screen "Dev_DO_2" 800x480, template "Settings"
   TextField "Text field_4" at 134,11 size 130x26; Text 'выход 1'
   TextField "Text field_5" at 286,11 size 130x26; Text 'выход 2'
   TextField "Text field_29" at 438,11 size 130x26; Text 'выход 3'
   TextField "Text field_33" at 590,11 size 130x26; Text 'выход 4'
   TextField "Text field_17" at 134,283 size 130x26; Text 'выход 9'
   TextField "Text field_25" at 286,283 size 130x26; Text 'выход 10'
   TextField "Text field_9" at 134,147 size 130x26; Text 'выход 5'
   TextField "Text field_13" at 286,147 size 130x26; Text 'выход 6'
   TextField "Text field_21" at 438,147 size 130x26; Text 'выход 7'
   TextField "Text field_41" at 590,147 size 130x26; Text 'выход 8'
   TextField "Text field_37" at 590,283 size 130x26; Text 'выход 12'
   Button "Button_2" at 134,40 size 130x22; TextOff 'Авто'; Authorization "Operate"; TextList "Hand"
      on Click: InvertBit("DOx_Hand_x_1")
      Appearance <- "DOx_Hand_x_1"
      ProcessValue <- "DOx_Hand_x_1"
   Button "Button_13" at 134,65 size 60x20; TextOff 'Вкл'; Authorization "Operate"
      on Click: SetBit("DOx_Start_M_x_1")
      Appearance <- "DOx_Start_M_x_1"
   Button "Button_26" at 244,89 size 20x20; TextOff 'Text'; Authorization "User administration"; PictureList "ok_green"
      on Click: InvertBit("DOx_Inverse_x_1")
      ProcessValue <- "DOx_Inverse_x_1"
   TextField "Text field_1" at 133,85 size 91x23; Text 'Инверсия:'
   IOField "I/O field_1" at 176,109 size 30x24; Authorization "Developer"; FormatPattern 99
      ProcessValue <- "DOx_ADDR_Byte_x_1"
   IOField "I/O field_2" at 216,109 size 20x24; Authorization "Developer"; FormatPattern 9
      ProcessValue <- "DOx_ADDR_Bit_x_1"
   TextField "Text field_2" at 158,109 size 20x23; Text 'Q'
   TextField "Text field_3" at 205,109 size 13x23; Text '.'
   Button "Button_1" at 286,40 size 130x22; TextOff 'Авто'; Authorization "Operate"; TextList "Hand"
      on Click: InvertBit("DOx_Hand_x_2")
      Appearance <- "DOx_Hand_x_2"
      ProcessValue <- "DOx_Hand_x_2"
   Button "Button_5" at 286,65 size 60x20; TextOff 'Вкл'; Authorization "Operate"
      on Click: SetBit("DOx_Start_M_x_2")
      Appearance <- "DOx_Start_M_x_2"
   Button "Button_6" at 396,89 size 20x20; TextOff 'Text'; PictureList "ok_green"; Authorization "User administration"
      on Click: InvertBit("DOx_Inverse_x_2")
      ProcessValue <- "DOx_Inverse_x_2"
   TextField "Text field_6" at 285,85 size 91x23; Text 'Инверсия:'
   IOField "I/O field_3" at 328,109 size 30x24; Authorization "Developer"; FormatPattern 99
      ProcessValue <- "DOx_ADDR_Byte_x_2"
   IOField "I/O field_4" at 368,109 size 20x24; Authorization "Developer"; FormatPattern 9
      ProcessValue <- "DOx_ADDR_Bit_x_2"
   TextField "Text field_7" at 310,109 size 20x23; Text 'Q'
   TextField "Text field_8" at 357,109 size 13x23; Text '.'
   Button "Button_29" at 438,40 size 130x22; TextOff 'Авто'; Authorization "Operate"; TextList "Hand"
      on Click: InvertBit("DOx_Hand_x_3")
      Appearance <- "DOx_Hand_x_3"
      ProcessValue <- "DOx_Hand_x_3"
   Button "Button_31" at 438,65 size 60x20; TextOff 'Вкл'; Authorization "Operate"
      on Click: SetBit("DOx_Start_M_x_3")
      Appearance <- "DOx_Start_M_x_3"
   Button "Button_32" at 548,89 size 20x20; TextOff 'Text'; PictureList "ok_green"; Authorization "User administration"
      on Click: InvertBit("DOx_Inverse_x_3")
      ProcessValue <- "DOx_Inverse_x_3"
   TextField "Text field_30" at 437,85 size 91x23; Text 'Инверсия:'
   IOField "I/O field_15" at 480,109 size 30x24; Authorization "Developer"; FormatPattern 99
      ProcessValue <- "DOx_ADDR_Byte_x_3"
   IOField "I/O field_16" at 520,109 size 20x24; Authorization "Developer"; FormatPattern 9
      ProcessValue <- "DOx_ADDR_Bit_x_3"
   TextField "Text field_31" at 462,109 size 20x23; Text 'Q'
   TextField "Text field_32" at 509,109 size 13x23; Text '.'
   Button "Button_33" at 590,40 size 130x22; TextOff 'Авто'; Authorization "Operate"; TextList "Hand"
      on Click: InvertBit("DOx_Hand_x_4")
      Appearance <- "DOx_Hand_x_4"
      ProcessValue <- "DOx_Hand_x_4"
   Button "Button_35" at 590,65 size 60x20; TextOff 'Вкл'; Authorization "Operate"
      on Click: SetBit("DOx_Start_M_x_4")
      Appearance <- "DOx_Start_M_x_4"
   Button "Button_36" at 700,89 size 20x20; TextOff 'Text'; PictureList "ok_green"; Authorization "User administration"
      on Click: InvertBit("DOx_Inverse_x_4")
      ProcessValue <- "DOx_Inverse_x_4"
   TextField "Text field_34" at 589,85 size 91x23; Text 'Инверсия:'
   IOField "I/O field_17" at 632,109 size 30x24; Authorization "Developer"; FormatPattern 99
      ProcessValue <- "DOx_ADDR_Byte_x_4"
   IOField "I/O field_18" at 672,109 size 20x24; Authorization "Developer"; FormatPattern 9
      ProcessValue <- "DOx_ADDR_Bit_x_4"
   TextField "Text field_35" at 614,109 size 20x23; Text 'Q'
   TextField "Text field_36" at 661,109 size 13x23; Text '.'
   Button "Button_7" at 134,176 size 130x22; TextOff 'Авто'; Authorization "Operate"; TextList "Hand"
      on Click: InvertBit("DOx_Hand_x_5")
      Appearance <- "DOx_Hand_x_5"
      ProcessValue <- "DOx_Hand_x_5"
   Button "Button_9" at 134,201 size 60x20; TextOff 'Вкл'; Authorization "Operate"
      on Click: SetBit("DOx_Start_M_x_5")
      Appearance <- "DOx_Start_M_x_5"
   Button "Button_10" at 244,225 size 20x20; TextOff 'Text'; PictureList "ok_green"; Authorization "User administration"
      on Click: InvertBit("DOx_Inverse_x_5")
      ProcessValue <- "DOx_Inverse_x_5"
   TextField "Text field_10" at 133,221 size 91x23; Text 'Инверсия:'
   IOField "I/O field_5" at 176,245 size 30x24; Authorization "Developer"; FormatPattern 99
      ProcessValue <- "DOx_ADDR_Byte_x_5"
   IOField "I/O field_6" at 216,245 size 20x24; Authorization "Developer"; FormatPattern 9
      ProcessValue <- "DOx_ADDR_Bit_x_5"
   TextField "Text field_11" at 158,245 size 20x23; Text 'Q'
   TextField "Text field_12" at 205,245 size 13x23; Text '.'
   Button "Button_11" at 286,176 size 130x22; TextOff 'Авто'; Authorization "Operate"; TextList "Hand"
      on Click: InvertBit("DOx_Hand_x_6")
      Appearance <- "DOx_Hand_x_6"
      ProcessValue <- "DOx_Hand_x_6"
   Button "Button_14" at 286,201 size 60x20; TextOff 'Вкл'; Authorization "Operate"
      on Click: SetBit("DOx_Start_M_x_6")
      Appearance <- "DOx_Start_M_x_6"
   Button "Button_15" at 396,225 size 20x20; TextOff 'Text'; Authorization "User administration"; PictureList "ok_green"
      on Click: InvertBit("DOx_Inverse_x_6")
      ProcessValue <- "DOx_Inverse_x_6"
   TextField "Text field_14" at 285,221 size 91x23; Text 'Инверсия:'
   IOField "I/O field_7" at 328,245 size 30x24; Authorization "Developer"; FormatPattern 99
      ProcessValue <- "DOx_ADDR_Byte_x_6"
   IOField "I/O field_8" at 368,245 size 20x24; Authorization "Developer"; FormatPattern 9
      ProcessValue <- "DOx_ADDR_Bit_x_6"
   TextField "Text field_15" at 310,245 size 20x23; Text 'Q'
   TextField "Text field_16" at 357,245 size 13x23; Text '.'
   Button "Button_20" at 438,176 size 130x22; TextOff 'Авто'; Authorization "Operate"; TextList "Hand"
      on Click: InvertBit("DOx_Hand_x_7")
      Appearance <- "DOx_Hand_x_7"
      ProcessValue <- "DOx_Hand_x_7"
   Button "Button_22" at 438,201 size 60x20; TextOff 'Вкл'; Authorization "Operate"
      on Click: SetBit("DOx_Start_M_x_7")
      Appearance <- "DOx_Start_M_x_7"
   Button "Button_23" at 548,225 size 20x20; TextOff 'Text'; Authorization "User administration"; PictureList "ok_green"
      on Click: InvertBit("DOx_Inverse_x_7")
      ProcessValue <- "DOx_Inverse_x_7"
   TextField "Text field_22" at 437,221 size 91x23; Text 'Инверсия:'
   IOField "I/O field_11" at 480,245 size 30x24; Authorization "Developer"; FormatPattern 99
      ProcessValue <- "DOx_ADDR_Byte_x_7"
   IOField "I/O field_12" at 520,245 size 20x24; Authorization "Developer"; FormatPattern 9
      ProcessValue <- "DOx_ADDR_Bit_x_7"
   TextField "Text field_23" at 462,245 size 20x23; Text 'Q'
   TextField "Text field_24" at 509,245 size 13x23; Text '.'
   Button "Button_41" at 590,176 size 130x22; TextOff 'Авто'; Authorization "Operate"; TextList "Hand"
      on Click: InvertBit("DOx_Hand_x_8")
      Appearance <- "DOx_Hand_x_8"
      ProcessValue <- "DOx_Hand_x_8"
   Button "Button_43" at 590,201 size 60x20; TextOff 'Вкл'; Authorization "Operate"
      on Click: SetBit("DOx_Start_M_x_8")
      Appearance <- "DOx_Start_M_x_8"
   Button "Button_44" at 700,225 size 20x20; TextOff 'Text'; Authorization "User administration"; PictureList "ok_green"
      on Click: InvertBit("DOx_Inverse_x_8")
      ProcessValue <- "DOx_Inverse_x_8"
   TextField "Text field_42" at 589,221 size 91x23; Text 'Инверсия:'
   IOField "I/O field_21" at 632,245 size 30x24; Authorization "Developer"; FormatPattern 99
      ProcessValue <- "DOx_ADDR_Byte_x_8"
   IOField "I/O field_22" at 672,245 size 20x24; Authorization "Developer"; FormatPattern 9
      ProcessValue <- "DOx_ADDR_Bit_x_8"
   TextField "Text field_43" at 614,245 size 20x23; Text 'Q'
   TextField "Text field_44" at 661,245 size 13x23; Text '.'
   Button "Button_24" at 134,312 size 130x22; TextOff 'Авто'; Authorization "Operate"; TextList "Hand"
      on Click: InvertBit("DOx_Hand_x_9")
      Appearance <- "DOx_Hand_x_9"
      ProcessValue <- "DOx_Hand_x_9"
   Button "Button_27" at 134,337 size 60x20; TextOff 'Вкл'; Authorization "Operate"
      on Click: SetBit("DOx_Start_M_x_9")
      Appearance <- "DOx_Start_M_x_9"
   Button "Button_28" at 244,361 size 20x20; TextOff 'Text'; PictureList "ok_green"; Authorization "User administration"
      on Click: InvertBit("DOx_Inverse_x_9")
      ProcessValue <- "DOx_Inverse_x_9"
   TextField "Text field_18" at 133,357 size 91x23; Text 'Инверсия:'
   IOField "I/O field_9" at 176,381 size 30x24; Authorization "Developer"; FormatPattern 99
      ProcessValue <- "DOx_ADDR_Byte_x_9"
   IOField "I/O field_10" at 216,381 size 20x24; Authorization "Developer"; FormatPattern 9
      ProcessValue <- "DOx_ADDR_Bit_x_9"
   TextField "Text field_19" at 158,381 size 20x23; Text 'Q'
   TextField "Text field_20" at 205,381 size 13x23; Text '.'
   Button "Button_37" at 286,312 size 130x22; TextOff 'Авто'; Authorization "Operate"; TextList "Hand"
      on Click: InvertBit("DOx_Hand_x_10")
      Appearance <- "DOx_Hand_x_10"
      ProcessValue <- "DOx_Hand_x_10"
   Button "Button_39" at 286,337 size 60x20; TextOff 'Вкл'; Authorization "Operate"
      on Click: SetBit("DOx_Start_M_x_10")
      Appearance <- "DOx_Start_M_x_10"
   Button "Button_40" at 396,361 size 20x20; TextOff 'Text'; Authorization "User administration"; PictureList "ok_green"
      on Click: InvertBit("DOx_Inverse_x_10")
      ProcessValue <- "DOx_Inverse_x_10"
   TextField "Text field_26" at 285,357 size 91x23; Text 'Инверсия:'
   IOField "I/O field_13" at 328,381 size 30x24; Authorization "Developer"; FormatPattern 99
      ProcessValue <- "DOx_ADDR_Byte_x_10"
   IOField "I/O field_14" at 368,381 size 20x24; Authorization "Developer"; FormatPattern 9
      ProcessValue <- "DOx_ADDR_Bit_x_10"
   TextField "Text field_27" at 310,381 size 20x23; Text 'Q'
   TextField "Text field_28" at 357,381 size 13x23; Text '.'
   Button "Button_48" at 590,312 size 130x22; TextOff 'Авто'; Authorization "Operate"; TextList "Hand"
      on Click: InvertBit("DOx_Hand_x_12")
      Appearance <- "DOx_Hand_x_12"
      ProcessValue <- "DOx_Hand_x_12"
   Button "Button_50" at 590,337 size 60x20; TextOff 'Вкл'; Authorization "Operate"
      on Click: SetBit("DOx_Start_M_x_12")
      Appearance <- "DOx_Start_M_x_12"
   Button "Button_51" at 700,361 size 20x20; TextOff 'Text'; Authorization "User administration"; PictureList "ok_green"
      on Click: InvertBit("DOx_Inverse_x_12")
      ProcessValue <- "DOx_Inverse_x_12"
   TextField "Text field_45" at 589,357 size 91x23; Text 'Инверсия:'
   IOField "I/O field_23" at 632,381 size 30x24; Authorization "Developer"; FormatPattern 99
      ProcessValue <- "DOx_ADDR_Byte_x_12"
   IOField "I/O field_24" at 672,381 size 20x24; Authorization "Developer"; FormatPattern 9
      ProcessValue <- "DOx_ADDR_Bit_x_12"
   TextField "Text field_46" at 614,381 size 20x23; Text 'Q'
   TextField "Text field_47" at 661,381 size 13x23; Text '.'
   TextField "Text field_38" at 438,283 size 130x26; Text 'выход 11'
   Button "Button_45" at 438,312 size 130x22; TextOff 'Авто'; Authorization "Operate"; TextList "Hand"
      on Click: InvertBit("DOx_Hand_x_11")
      Appearance <- "DOx_Hand_x_11"
      ProcessValue <- "DOx_Hand_x_11"
   Button "Button_47" at 438,337 size 60x20; TextOff 'Вкл'; Authorization "Operate"
      on Click: SetBit("DOx_Start_M_x_11")
      Appearance <- "DOx_Start_M_x_11"
   Button "Button_52" at 548,361 size 20x20; TextOff 'Text'; PictureList "ok_green"; Authorization "User administration"
      on Click: InvertBit("DOx_Inverse_x_11")
      ProcessValue <- "DOx_Inverse_x_11"
   TextField "Text field_39" at 437,357 size 91x23; Text 'Инверсия:'
   IOField "I/O field_19" at 480,381 size 30x24; Authorization "Developer"; FormatPattern 99
      ProcessValue <- "DOx_ADDR_Byte_x_11"
   IOField "I/O field_20" at 520,381 size 20x24; Authorization "Developer"; FormatPattern 9
      ProcessValue <- "DOx_ADDR_Bit_x_11"
   TextField "Text field_40" at 462,381 size 20x23; Text 'Q'
   TextField "Text field_48" at 509,381 size 13x23; Text '.'
   Button "Button_16" at 128,440 size 75x30; TextOff 'Стр.1'; Authorization "Operate"
      on Click: SetTag("DOx", 210); ActivateScreen("Dev_DI_1", 0)
      Visibility <- "Support_DB_All_DOs"
      Appearance <- "DOx"
   Button "Button_17" at 233,440 size 75x30; TextOff 'Стр.2'; Authorization "Operate"
      on Click: SetTag("DOx", 211); ActivateScreen("Dev_DI_2", 0)
      Visibility <- "Support_DB_All_DOs"
      Appearance <- "DOx"
   Button "Button_18" at 338,440 size 75x30; TextOff 'Стр.3'; Authorization "Operate"
      on Click: SetTag("DOx", 212); ActivateScreen("Dev_DI_3", 0)
      Visibility <- "Support_DB_All_DOs"
      Appearance <- "DOx"
   Button "Button_19" at 444,440 size 75x30; TextOff 'Стр.4'; Authorization "Operate"
      on Click: SetTag("DOx", 213); ActivateScreen("Dev_DI_4", 0)
      Visibility <- "Support_DB_All_DOs"
      Appearance <- "DOx"
   Button "Button_53" at 549,440 size 75x30; TextOff 'Стр.5'; Authorization "Operate"
      on Click: SetTag("DOx", 214); ActivateScreen("Dev_DI_5", 0)
      Visibility <- "Support_DB_All_DOs"
      Appearance <- "DOx"
   Button "Button_54" at 655,440 size 75x30; TextOff 'Стр.6'; Authorization "Operate"
      on Click: SetTag("DOx", 215); ActivateScreen("Dev_DI_6", 0)
      Visibility <- "Support_DB_All_DOs"
      Appearance <- "DOx"
   Button "Button_3" at 204,65 size 60x20; TextOff 'Выкл'; Authorization "Operate"
      on Click: ResetBit("DOx_Start_M_x_1")
      Appearance <- "DOx_Start_M_x_1"
   Button "Button_4" at 356,65 size 60x20; TextOff 'Выкл'; Authorization "Operate"
      on Click: ResetBit("DOx_Start_M_x_2")
      Appearance <- "DOx_Start_M_x_2"
   Button "Button_30" at 508,65 size 60x20; TextOff 'Выкл'; Authorization "Operate"
      on Click: ResetBit("DOx_Start_M_x_3")
      Appearance <- "DOx_Start_M_x_3"
   Button "Button_34" at 660,65 size 60x20; TextOff 'Выкл'; Authorization "Operate"
      on Click: ResetBit("DOx_Start_M_x_4")
      Appearance <- "DOx_Start_M_x_4"
   Button "Button_8" at 204,201 size 60x20; TextOff 'Выкл'; Authorization "Operate"
      on Click: ResetBit("DOx_Start_M_x_5")
      Appearance <- "DOx_Start_M_x_5"
   Button "Button_12" at 356,201 size 60x20; TextOff 'Выкл'; Authorization "Operate"
      on Click: ResetBit("DOx_Start_M_x_6")
      Appearance <- "DOx_Start_M_x_6"
   Button "Button_21" at 508,201 size 60x20; TextOff 'Выкл'; Authorization "Operate"
      on Click: ResetBit("DOx_Start_M_x_7")
      Appearance <- "DOx_Start_M_x_7"
   Button "Button_42" at 660,201 size 60x20; TextOff 'Выкл'; Authorization "Operate"
      on Click: ResetBit("DOx_Start_M_x_8")
      Appearance <- "DOx_Start_M_x_8"
   Button "Button_25" at 204,337 size 60x20; TextOff 'Выкл'; Authorization "Operate"
      on Click: ResetBit("DOx_Start_M_x_9")
      Appearance <- "DOx_Start_M_x_9"
   Button "Button_38" at 356,337 size 60x20; TextOff 'Выкл'; Authorization "Operate"
      on Click: ResetBit("DOx_Start_M_x_10")
      Appearance <- "DOx_Start_M_x_10"
   Button "Button_49" at 660,337 size 60x20; TextOff 'Выкл'; Authorization "Operate"
      on Click: ResetBit("DOx_Start_M_x_12")
      Appearance <- "DOx_Start_M_x_12"
   Button "Button_46" at 508,337 size 60x20; TextOff 'Выкл'; Authorization "Operate"
      on Click: ResetBit("DOx_Start_M_x_11")
      Appearance <- "DOx_Start_M_x_11"

screen "Dev_DO_3" 800x480, template "Settings"
   TextField "Text field_4" at 134,11 size 130x26; Text 'выход 1'
   TextField "Text field_5" at 286,11 size 130x26; Text 'выход 2'
   TextField "Text field_29" at 438,11 size 130x26; Text 'выход 3'
   TextField "Text field_33" at 590,11 size 130x26; Text 'выход 4'
   TextField "Text field_17" at 134,283 size 130x26; Text 'выход 9'
   TextField "Text field_25" at 286,283 size 130x26; Text 'выход 10'
   TextField "Text field_9" at 134,147 size 130x26; Text 'выход 5'
   TextField "Text field_13" at 286,147 size 130x26; Text 'выход 6'
   TextField "Text field_21" at 438,147 size 130x26; Text 'выход 7'
   TextField "Text field_41" at 590,147 size 130x26; Text 'выход 8'
   TextField "Text field_37" at 590,283 size 130x26; Text 'выход 12'
   Button "Button_2" at 134,40 size 130x22; TextOff 'Авто'; Authorization "Operate"; TextList "Hand"
      on Click: InvertBit("DOx_Hand_x_1")
      Appearance <- "DOx_Hand_x_1"
      ProcessValue <- "DOx_Hand_x_1"
   Button "Button_13" at 134,65 size 60x20; TextOff 'Вкл'; Authorization "Operate"
      on Click: SetBit("DOx_Start_M_x_1")
      Appearance <- "DOx_Start_M_x_1"
   Button "Button_26" at 244,89 size 20x20; TextOff 'Text'; Authorization "User administration"; PictureList "ok_green"
      on Click: InvertBit("DOx_Inverse_x_1")
      ProcessValue <- "DOx_Inverse_x_1"
   TextField "Text field_1" at 133,85 size 91x23; Text 'Инверсия:'
   IOField "I/O field_1" at 176,109 size 30x24; Authorization "Developer"; FormatPattern 99
      ProcessValue <- "DOx_ADDR_Byte_x_1"
   IOField "I/O field_2" at 216,109 size 20x24; Authorization "Developer"; FormatPattern 9
      ProcessValue <- "DOx_ADDR_Bit_x_1"
   TextField "Text field_2" at 158,109 size 20x23; Text 'Q'
   TextField "Text field_3" at 205,109 size 13x23; Text '.'
   Button "Button_1" at 286,40 size 130x22; TextOff 'Авто'; Authorization "Operate"; TextList "Hand"
      on Click: InvertBit("DOx_Hand_x_2")
      Appearance <- "DOx_Hand_x_2"
      ProcessValue <- "DOx_Hand_x_2"
   Button "Button_5" at 286,65 size 60x20; TextOff 'Вкл'; Authorization "Operate"
      on Click: SetBit("DOx_Start_M_x_2")
      Appearance <- "DOx_Start_M_x_2"
   Button "Button_6" at 396,89 size 20x20; TextOff 'Text'; PictureList "ok_green"; Authorization "User administration"
      on Click: InvertBit("DOx_Inverse_x_2")
      ProcessValue <- "DOx_Inverse_x_2"
   TextField "Text field_6" at 285,85 size 91x23; Text 'Инверсия:'
   IOField "I/O field_3" at 328,109 size 30x24; Authorization "Developer"; FormatPattern 99
      ProcessValue <- "DOx_ADDR_Byte_x_2"
   IOField "I/O field_4" at 368,109 size 20x24; Authorization "Developer"; FormatPattern 9
      ProcessValue <- "DOx_ADDR_Bit_x_2"
   TextField "Text field_7" at 310,109 size 20x23; Text 'Q'
   TextField "Text field_8" at 357,109 size 13x23; Text '.'
   Button "Button_29" at 438,40 size 130x22; TextOff 'Авто'; Authorization "Operate"; TextList "Hand"
      on Click: InvertBit("DOx_Hand_x_3")
      Appearance <- "DOx_Hand_x_3"
      ProcessValue <- "DOx_Hand_x_3"
   Button "Button_31" at 438,65 size 60x20; TextOff 'Вкл'; Authorization "Operate"
      on Click: SetBit("DOx_Start_M_x_3")
      Appearance <- "DOx_Start_M_x_3"
   Button "Button_32" at 548,89 size 20x20; TextOff 'Text'; PictureList "ok_green"; Authorization "User administration"
      on Click: InvertBit("DOx_Inverse_x_3")
      ProcessValue <- "DOx_Inverse_x_3"
   TextField "Text field_30" at 437,85 size 91x23; Text 'Инверсия:'
   IOField "I/O field_15" at 480,109 size 30x24; Authorization "Developer"; FormatPattern 99
      ProcessValue <- "DOx_ADDR_Byte_x_3"
   IOField "I/O field_16" at 520,109 size 20x24; Authorization "Developer"; FormatPattern 9
      ProcessValue <- "DOx_ADDR_Bit_x_3"
   TextField "Text field_31" at 462,109 size 20x23; Text 'Q'
   TextField "Text field_32" at 509,109 size 13x23; Text '.'
   Button "Button_33" at 590,40 size 130x22; TextOff 'Авто'; Authorization "Operate"; TextList "Hand"
      on Click: InvertBit("DOx_Hand_x_4")
      Appearance <- "DOx_Hand_x_4"
      ProcessValue <- "DOx_Hand_x_4"
   Button "Button_35" at 590,65 size 60x20; TextOff 'Вкл'; Authorization "Operate"
      on Click: SetBit("DOx_Start_M_x_4")
      Appearance <- "DOx_Start_M_x_4"
   Button "Button_36" at 700,89 size 20x20; TextOff 'Text'; PictureList "ok_green"; Authorization "User administration"
      on Click: InvertBit("DOx_Inverse_x_4")
      ProcessValue <- "DOx_Inverse_x_4"
   TextField "Text field_34" at 589,85 size 91x23; Text 'Инверсия:'
   IOField "I/O field_17" at 632,109 size 30x24; Authorization "Developer"; FormatPattern 99
      ProcessValue <- "DOx_ADDR_Byte_x_4"
   IOField "I/O field_18" at 672,109 size 20x24; Authorization "Developer"; FormatPattern 9
      ProcessValue <- "DOx_ADDR_Bit_x_4"
   TextField "Text field_35" at 614,109 size 20x23; Text 'Q'
   TextField "Text field_36" at 661,109 size 13x23; Text '.'
   Button "Button_7" at 134,176 size 130x22; TextOff 'Авто'; Authorization "Operate"; TextList "Hand"
      on Click: InvertBit("DOx_Hand_x_5")
      Appearance <- "DOx_Hand_x_5"
      ProcessValue <- "DOx_Hand_x_5"
   Button "Button_9" at 134,201 size 60x20; TextOff 'Вкл'; Authorization "Operate"
      on Click: SetBit("DOx_Start_M_x_5")
      Appearance <- "DOx_Start_M_x_5"
   Button "Button_10" at 244,225 size 20x20; TextOff 'Text'; PictureList "ok_green"; Authorization "User administration"
      on Click: InvertBit("DOx_Inverse_x_5")
      ProcessValue <- "DOx_Inverse_x_5"
   TextField "Text field_10" at 133,221 size 91x23; Text 'Инверсия:'
   IOField "I/O field_5" at 176,245 size 30x24; Authorization "Developer"; FormatPattern 99
      ProcessValue <- "DOx_ADDR_Byte_x_5"
   IOField "I/O field_6" at 216,245 size 20x24; Authorization "Developer"; FormatPattern 9
      ProcessValue <- "DOx_ADDR_Bit_x_5"
   TextField "Text field_11" at 158,245 size 20x23; Text 'Q'
   TextField "Text field_12" at 205,245 size 13x23; Text '.'
   Button "Button_11" at 286,176 size 130x22; TextOff 'Авто'; Authorization "Operate"; TextList "Hand"
      on Click: InvertBit("DOx_Hand_x_6")
      Appearance <- "DOx_Hand_x_6"
      ProcessValue <- "DOx_Hand_x_6"
   Button "Button_14" at 286,201 size 60x20; TextOff 'Вкл'; Authorization "Operate"
      on Click: SetBit("DOx_Start_M_x_6")
      Appearance <- "DOx_Start_M_x_6"
   Button "Button_15" at 396,225 size 20x20; TextOff 'Text'; Authorization "User administration"; PictureList "ok_green"
      on Click: InvertBit("DOx_Inverse_x_6")
      ProcessValue <- "DOx_Inverse_x_6"
   TextField "Text field_14" at 285,221 size 91x23; Text 'Инверсия:'
   IOField "I/O field_7" at 328,245 size 30x24; Authorization "Developer"; FormatPattern 99
      ProcessValue <- "DOx_ADDR_Byte_x_6"
   IOField "I/O field_8" at 368,245 size 20x24; Authorization "Developer"; FormatPattern 9
      ProcessValue <- "DOx_ADDR_Bit_x_6"
   TextField "Text field_15" at 310,245 size 20x23; Text 'Q'
   TextField "Text field_16" at 357,245 size 13x23; Text '.'
   Button "Button_20" at 438,176 size 130x22; TextOff 'Авто'; Authorization "Operate"; TextList "Hand"
      on Click: InvertBit("DOx_Hand_x_7")
      Appearance <- "DOx_Hand_x_7"
      ProcessValue <- "DOx_Hand_x_7"
   Button "Button_22" at 438,201 size 60x20; TextOff 'Вкл'; Authorization "Operate"
      on Click: SetBit("DOx_Start_M_x_7")
      Appearance <- "DOx_Start_M_x_7"
   Button "Button_23" at 548,225 size 20x20; TextOff 'Text'; Authorization "User administration"; PictureList "ok_green"
      on Click: InvertBit("DOx_Inverse_x_7")
      ProcessValue <- "DOx_Inverse_x_7"
   TextField "Text field_22" at 437,221 size 91x23; Text 'Инверсия:'
   IOField "I/O field_11" at 480,245 size 30x24; Authorization "Developer"; FormatPattern 99
      ProcessValue <- "DOx_ADDR_Byte_x_7"
   IOField "I/O field_12" at 520,245 size 20x24; Authorization "Developer"; FormatPattern 9
      ProcessValue <- "DOx_ADDR_Bit_x_7"
   TextField "Text field_23" at 462,245 size 20x23; Text 'Q'
   TextField "Text field_24" at 509,245 size 13x23; Text '.'
   Button "Button_41" at 590,176 size 130x22; TextOff 'Авто'; Authorization "Operate"; TextList "Hand"
      on Click: InvertBit("DOx_Hand_x_8")
      Appearance <- "DOx_Hand_x_8"
      ProcessValue <- "DOx_Hand_x_8"
   Button "Button_43" at 590,201 size 60x20; TextOff 'Вкл'; Authorization "Operate"
      on Click: SetBit("DOx_Start_M_x_8")
      Appearance <- "DOx_Start_M_x_8"
   Button "Button_44" at 700,225 size 20x20; TextOff 'Text'; Authorization "User administration"; PictureList "ok_green"
      on Click: InvertBit("DOx_Inverse_x_8")
      ProcessValue <- "DOx_Inverse_x_8"
   TextField "Text field_42" at 589,221 size 91x23; Text 'Инверсия:'
   IOField "I/O field_21" at 632,245 size 30x24; Authorization "Developer"; FormatPattern 99
      ProcessValue <- "DOx_ADDR_Byte_x_8"
   IOField "I/O field_22" at 672,245 size 20x24; Authorization "Developer"; FormatPattern 9
      ProcessValue <- "DOx_ADDR_Bit_x_8"
   TextField "Text field_43" at 614,245 size 20x23; Text 'Q'
   TextField "Text field_44" at 661,245 size 13x23; Text '.'
   Button "Button_24" at 134,312 size 130x22; TextOff 'Авто'; Authorization "Operate"; TextList "Hand"
      on Click: InvertBit("DOx_Hand_x_9")
      Appearance <- "DOx_Hand_x_9"
      ProcessValue <- "DOx_Hand_x_9"
   Button "Button_27" at 134,337 size 60x20; TextOff 'Вкл'; Authorization "Operate"
      on Click: SetBit("DOx_Start_M_x_9")
      Appearance <- "DOx_Start_M_x_9"
   Button "Button_28" at 244,361 size 20x20; TextOff 'Text'; PictureList "ok_green"; Authorization "User administration"
      on Click: InvertBit("DOx_Inverse_x_9")
      ProcessValue <- "DOx_Inverse_x_9"
   TextField "Text field_18" at 133,357 size 91x23; Text 'Инверсия:'
   IOField "I/O field_9" at 176,381 size 30x24; Authorization "Developer"; FormatPattern 99
      ProcessValue <- "DOx_ADDR_Byte_x_9"
   IOField "I/O field_10" at 216,381 size 20x24; Authorization "Developer"; FormatPattern 9
      ProcessValue <- "DOx_ADDR_Bit_x_9"
   TextField "Text field_19" at 158,381 size 20x23; Text 'Q'
   TextField "Text field_20" at 205,381 size 13x23; Text '.'
   Button "Button_37" at 286,312 size 130x22; TextOff 'Авто'; Authorization "Operate"; TextList "Hand"
      on Click: InvertBit("DOx_Hand_x_10")
      Appearance <- "DOx_Hand_x_10"
      ProcessValue <- "DOx_Hand_x_10"
   Button "Button_39" at 286,337 size 60x20; TextOff 'Вкл'; Authorization "Operate"
      on Click: SetBit("DOx_Start_M_x_10")
      Appearance <- "DOx_Start_M_x_10"
   Button "Button_40" at 396,361 size 20x20; TextOff 'Text'; Authorization "User administration"; PictureList "ok_green"
      on Click: InvertBit("DOx_Inverse_x_10")
      ProcessValue <- "DOx_Inverse_x_10"
   TextField "Text field_26" at 285,357 size 91x23; Text 'Инверсия:'
   IOField "I/O field_13" at 328,381 size 30x24; Authorization "Developer"; FormatPattern 99
      ProcessValue <- "DOx_ADDR_Byte_x_10"
   IOField "I/O field_14" at 368,381 size 20x24; Authorization "Developer"; FormatPattern 9
      ProcessValue <- "DOx_ADDR_Bit_x_10"
   TextField "Text field_27" at 310,381 size 20x23; Text 'Q'
   TextField "Text field_28" at 357,381 size 13x23; Text '.'
   Button "Button_48" at 590,312 size 130x22; TextOff 'Авто'; Authorization "Operate"; TextList "Hand"
      on Click: InvertBit("DOx_Hand_x_12")
      Appearance <- "DOx_Hand_x_12"
      ProcessValue <- "DOx_Hand_x_12"
   Button "Button_50" at 590,337 size 60x20; TextOff 'Вкл'; Authorization "Operate"
      on Click: SetBit("DOx_Start_M_x_12")
      Appearance <- "DOx_Start_M_x_12"
   Button "Button_51" at 700,361 size 20x20; TextOff 'Text'; Authorization "User administration"; PictureList "ok_green"
      on Click: InvertBit("DOx_Inverse_x_12")
      ProcessValue <- "DOx_Inverse_x_12"
   TextField "Text field_45" at 589,357 size 91x23; Text 'Инверсия:'
   IOField "I/O field_23" at 632,381 size 30x24; Authorization "Developer"; FormatPattern 99
      ProcessValue <- "DOx_ADDR_Byte_x_12"
   IOField "I/O field_24" at 672,381 size 20x24; Authorization "Developer"; FormatPattern 9
      ProcessValue <- "DOx_ADDR_Bit_x_12"
   TextField "Text field_46" at 614,381 size 20x23; Text 'Q'
   TextField "Text field_47" at 661,381 size 13x23; Text '.'
   TextField "Text field_38" at 438,283 size 130x26; Text 'выход 11'
   Button "Button_45" at 438,312 size 130x22; TextOff 'Авто'; Authorization "Operate"; TextList "Hand"
      on Click: InvertBit("DOx_Hand_x_11")
      Appearance <- "DOx_Hand_x_11"
      ProcessValue <- "DOx_Hand_x_11"
   Button "Button_47" at 438,337 size 60x20; TextOff 'Вкл'; Authorization "Operate"
      on Click: SetBit("DOx_Start_M_x_11")
      Appearance <- "DOx_Start_M_x_11"
   Button "Button_52" at 548,361 size 20x20; TextOff 'Text'; PictureList "ok_green"; Authorization "User administration"
      on Click: InvertBit("DOx_Inverse_x_11")
      ProcessValue <- "DOx_Inverse_x_11"
   TextField "Text field_39" at 437,357 size 91x23; Text 'Инверсия:'
   IOField "I/O field_19" at 480,381 size 30x24; Authorization "Developer"; FormatPattern 99
      ProcessValue <- "DOx_ADDR_Byte_x_11"
   IOField "I/O field_20" at 520,381 size 20x24; Authorization "Developer"; FormatPattern 9
      ProcessValue <- "DOx_ADDR_Bit_x_11"
   TextField "Text field_40" at 462,381 size 20x23; Text 'Q'
   TextField "Text field_48" at 509,381 size 13x23; Text '.'
   Button "Button_16" at 128,440 size 75x30; TextOff 'Стр.1'; Authorization "Operate"
      on Click: SetTag("DOx", 210); ActivateScreen("Dev_DI_1", 0)
      Visibility <- "Support_DB_All_DOs"
      Appearance <- "DOx"
   Button "Button_17" at 233,440 size 75x30; TextOff 'Стр.2'; Authorization "Operate"
      on Click: SetTag("DOx", 211); ActivateScreen("Dev_DI_2", 0)
      Visibility <- "Support_DB_All_DOs"
      Appearance <- "DOx"
   Button "Button_18" at 338,440 size 75x30; TextOff 'Стр.3'; Authorization "Operate"
      on Click: SetTag("DOx", 212); ActivateScreen("Dev_DI_3", 0)
      Visibility <- "Support_DB_All_DOs"
      Appearance <- "DOx"
   Button "Button_19" at 444,440 size 75x30; TextOff 'Стр.4'; Authorization "Operate"
      on Click: SetTag("DOx", 213); ActivateScreen("Dev_DI_4", 0)
      Visibility <- "Support_DB_All_DOs"
      Appearance <- "DOx"
   Button "Button_53" at 549,440 size 75x30; TextOff 'Стр.5'; Authorization "Operate"
      on Click: SetTag("DOx", 214); ActivateScreen("Dev_DI_5", 0)
      Visibility <- "Support_DB_All_DOs"
      Appearance <- "DOx"
   Button "Button_54" at 655,440 size 75x30; TextOff 'Стр.6'; Authorization "Operate"
      on Click: SetTag("DOx", 215); ActivateScreen("Dev_DI_6", 0)
      Visibility <- "Support_DB_All_DOs"
      Appearance <- "DOx"
   Button "Button_3" at 204,65 size 60x20; TextOff 'Выкл'; Authorization "Operate"
      on Click: ResetBit("DOx_Start_M_x_1")
      Appearance <- "DOx_Start_M_x_1"
   Button "Button_4" at 356,65 size 60x20; TextOff 'Выкл'; Authorization "Operate"
      on Click: ResetBit("DOx_Start_M_x_2")
      Appearance <- "DOx_Start_M_x_2"
   Button "Button_30" at 508,65 size 60x20; TextOff 'Выкл'; Authorization "Operate"
      on Click: ResetBit("DOx_Start_M_x_3")
      Appearance <- "DOx_Start_M_x_3"
   Button "Button_34" at 660,65 size 60x20; TextOff 'Выкл'; Authorization "Operate"
      on Click: ResetBit("DOx_Start_M_x_4")
      Appearance <- "DOx_Start_M_x_4"
   Button "Button_8" at 204,201 size 60x20; TextOff 'Выкл'; Authorization "Operate"
      on Click: ResetBit("DOx_Start_M_x_5")
      Appearance <- "DOx_Start_M_x_5"
   Button "Button_12" at 356,201 size 60x20; TextOff 'Выкл'; Authorization "Operate"
      on Click: ResetBit("DOx_Start_M_x_6")
      Appearance <- "DOx_Start_M_x_6"
   Button "Button_21" at 508,201 size 60x20; TextOff 'Выкл'; Authorization "Operate"
      on Click: ResetBit("DOx_Start_M_x_7")
      Appearance <- "DOx_Start_M_x_7"
   Button "Button_42" at 660,201 size 60x20; TextOff 'Выкл'; Authorization "Operate"
      on Click: ResetBit("DOx_Start_M_x_8")
      Appearance <- "DOx_Start_M_x_8"
   Button "Button_25" at 204,337 size 60x20; TextOff 'Выкл'; Authorization "Operate"
      on Click: ResetBit("DOx_Start_M_x_9")
      Appearance <- "DOx_Start_M_x_9"
   Button "Button_38" at 356,337 size 60x20; TextOff 'Выкл'; Authorization "Operate"
      on Click: ResetBit("DOx_Start_M_x_10")
      Appearance <- "DOx_Start_M_x_10"
   Button "Button_49" at 660,337 size 60x20; TextOff 'Выкл'; Authorization "Operate"
      on Click: ResetBit("DOx_Start_M_x_12")
      Appearance <- "DOx_Start_M_x_12"
   Button "Button_46" at 508,337 size 60x20; TextOff 'Выкл'; Authorization "Operate"
      on Click: ResetBit("DOx_Start_M_x_11")
      Appearance <- "DOx_Start_M_x_11"

screen "Dev_DO_4" 800x480, template "Settings"
   TextField "Text field_4" at 134,11 size 130x26; Text 'выход 1'
   TextField "Text field_5" at 286,11 size 130x26; Text 'выход 2'
   TextField "Text field_29" at 438,11 size 130x26; Text 'выход 3'
   TextField "Text field_33" at 590,11 size 130x26; Text 'выход 4'
   TextField "Text field_17" at 134,283 size 130x26; Text 'выход 9'
   TextField "Text field_25" at 286,283 size 130x26; Text 'выход 10'
   TextField "Text field_9" at 134,147 size 130x26; Text 'выход 5'
   TextField "Text field_13" at 286,147 size 130x26; Text 'выход 6'
   TextField "Text field_21" at 438,147 size 130x26; Text 'выход 7'
   TextField "Text field_41" at 590,147 size 130x26; Text 'выход 8'
   TextField "Text field_37" at 590,283 size 130x26; Text 'выход 12'
   Button "Button_2" at 134,40 size 130x22; TextOff 'Авто'; Authorization "Operate"; TextList "Hand"
      on Click: InvertBit("DOx_Hand_x_1")
      Appearance <- "DOx_Hand_x_1"
      ProcessValue <- "DOx_Hand_x_1"
   Button "Button_13" at 134,65 size 60x20; TextOff 'Вкл'; Authorization "Operate"
      on Click: SetBit("DOx_Start_M_x_1")
      Appearance <- "DOx_Start_M_x_1"
   Button "Button_26" at 244,89 size 20x20; TextOff 'Text'; Authorization "User administration"; PictureList "ok_green"
      on Click: InvertBit("DOx_Inverse_x_1")
      ProcessValue <- "DOx_Inverse_x_1"
   TextField "Text field_1" at 133,85 size 91x23; Text 'Инверсия:'
   IOField "I/O field_1" at 176,109 size 30x24; Authorization "Developer"; FormatPattern 99
      ProcessValue <- "DOx_ADDR_Byte_x_1"
   IOField "I/O field_2" at 216,109 size 20x24; Authorization "Developer"; FormatPattern 9
      ProcessValue <- "DOx_ADDR_Bit_x_1"
   TextField "Text field_2" at 158,109 size 20x23; Text 'Q'
   TextField "Text field_3" at 205,109 size 13x23; Text '.'
   Button "Button_1" at 286,40 size 130x22; TextOff 'Авто'; Authorization "Operate"; TextList "Hand"
      on Click: InvertBit("DOx_Hand_x_2")
      Appearance <- "DOx_Hand_x_2"
      ProcessValue <- "DOx_Hand_x_2"
   Button "Button_5" at 286,65 size 60x20; TextOff 'Вкл'; Authorization "Operate"
      on Click: SetBit("DOx_Start_M_x_2")
      Appearance <- "DOx_Start_M_x_2"
   Button "Button_6" at 396,89 size 20x20; TextOff 'Text'; PictureList "ok_green"; Authorization "User administration"
      on Click: InvertBit("DOx_Inverse_x_2")
      ProcessValue <- "DOx_Inverse_x_2"
   TextField "Text field_6" at 285,85 size 91x23; Text 'Инверсия:'
   IOField "I/O field_3" at 328,109 size 30x24; Authorization "Developer"; FormatPattern 99
      ProcessValue <- "DOx_ADDR_Byte_x_2"
   IOField "I/O field_4" at 368,109 size 20x24; Authorization "Developer"; FormatPattern 9
      ProcessValue <- "DOx_ADDR_Bit_x_2"
   TextField "Text field_7" at 310,109 size 20x23; Text 'Q'
   TextField "Text field_8" at 357,109 size 13x23; Text '.'
   Button "Button_29" at 438,40 size 130x22; TextOff 'Авто'; Authorization "Operate"; TextList "Hand"
      on Click: InvertBit("DOx_Hand_x_3")
      Appearance <- "DOx_Hand_x_3"
      ProcessValue <- "DOx_Hand_x_3"
   Button "Button_31" at 438,65 size 60x20; TextOff 'Вкл'; Authorization "Operate"
      on Click: SetBit("DOx_Start_M_x_3")
      Appearance <- "DOx_Start_M_x_3"
   Button "Button_32" at 548,89 size 20x20; TextOff 'Text'; PictureList "ok_green"; Authorization "User administration"
      on Click: InvertBit("DOx_Inverse_x_3")
      ProcessValue <- "DOx_Inverse_x_3"
   TextField "Text field_30" at 437,85 size 91x23; Text 'Инверсия:'
   IOField "I/O field_15" at 480,109 size 30x24; Authorization "Developer"; FormatPattern 99
      ProcessValue <- "DOx_ADDR_Byte_x_3"
   IOField "I/O field_16" at 520,109 size 20x24; Authorization "Developer"; FormatPattern 9
      ProcessValue <- "DOx_ADDR_Bit_x_3"
   TextField "Text field_31" at 462,109 size 20x23; Text 'Q'
   TextField "Text field_32" at 509,109 size 13x23; Text '.'
   Button "Button_33" at 590,40 size 130x22; TextOff 'Авто'; Authorization "Operate"; TextList "Hand"
      on Click: InvertBit("DOx_Hand_x_4")
      Appearance <- "DOx_Hand_x_4"
      ProcessValue <- "DOx_Hand_x_4"
   Button "Button_35" at 590,65 size 60x20; TextOff 'Вкл'; Authorization "Operate"
      on Click: SetBit("DOx_Start_M_x_4")
      Appearance <- "DOx_Start_M_x_4"
   Button "Button_36" at 700,89 size 20x20; TextOff 'Text'; PictureList "ok_green"; Authorization "User administration"
      on Click: InvertBit("DOx_Inverse_x_4")
      ProcessValue <- "DOx_Inverse_x_4"
   TextField "Text field_34" at 589,85 size 91x23; Text 'Инверсия:'
   IOField "I/O field_17" at 632,109 size 30x24; Authorization "Developer"; FormatPattern 99
      ProcessValue <- "DOx_ADDR_Byte_x_4"
   IOField "I/O field_18" at 672,109 size 20x24; Authorization "Developer"; FormatPattern 9
      ProcessValue <- "DOx_ADDR_Bit_x_4"
   TextField "Text field_35" at 614,109 size 20x23; Text 'Q'
   TextField "Text field_36" at 661,109 size 13x23; Text '.'
   Button "Button_7" at 134,176 size 130x22; TextOff 'Авто'; Authorization "Operate"; TextList "Hand"
      on Click: InvertBit("DOx_Hand_x_5")
      Appearance <- "DOx_Hand_x_5"
      ProcessValue <- "DOx_Hand_x_5"
   Button "Button_9" at 134,201 size 60x20; TextOff 'Вкл'; Authorization "Operate"
      on Click: SetBit("DOx_Start_M_x_5")
      Appearance <- "DOx_Start_M_x_5"
   Button "Button_10" at 244,225 size 20x20; TextOff 'Text'; PictureList "ok_green"; Authorization "User administration"
      on Click: InvertBit("DOx_Inverse_x_5")
      ProcessValue <- "DOx_Inverse_x_5"
   TextField "Text field_10" at 133,221 size 91x23; Text 'Инверсия:'
   IOField "I/O field_5" at 176,245 size 30x24; Authorization "Developer"; FormatPattern 99
      ProcessValue <- "DOx_ADDR_Byte_x_5"
   IOField "I/O field_6" at 216,245 size 20x24; Authorization "Developer"; FormatPattern 9
      ProcessValue <- "DOx_ADDR_Bit_x_5"
   TextField "Text field_11" at 158,245 size 20x23; Text 'Q'
   TextField "Text field_12" at 205,245 size 13x23; Text '.'
   Button "Button_11" at 286,176 size 130x22; TextOff 'Авто'; Authorization "Operate"; TextList "Hand"
      on Click: InvertBit("DOx_Hand_x_6")
      Appearance <- "DOx_Hand_x_6"
      ProcessValue <- "DOx_Hand_x_6"
   Button "Button_14" at 286,201 size 60x20; TextOff 'Вкл'; Authorization "Operate"
      on Click: SetBit("DOx_Start_M_x_6")
      Appearance <- "DOx_Start_M_x_6"
   Button "Button_15" at 396,225 size 20x20; TextOff 'Text'; Authorization "User administration"; PictureList "ok_green"
      on Click: InvertBit("DOx_Inverse_x_6")
      ProcessValue <- "DOx_Inverse_x_6"
   TextField "Text field_14" at 285,221 size 91x23; Text 'Инверсия:'
   IOField "I/O field_7" at 328,245 size 30x24; Authorization "Developer"; FormatPattern 99
      ProcessValue <- "DOx_ADDR_Byte_x_6"
   IOField "I/O field_8" at 368,245 size 20x24; Authorization "Developer"; FormatPattern 9
      ProcessValue <- "DOx_ADDR_Bit_x_6"
   TextField "Text field_15" at 310,245 size 20x23; Text 'Q'
   TextField "Text field_16" at 357,245 size 13x23; Text '.'
   Button "Button_20" at 438,176 size 130x22; TextOff 'Авто'; Authorization "Operate"; TextList "Hand"
      on Click: InvertBit("DOx_Hand_x_7")
      Appearance <- "DOx_Hand_x_7"
      ProcessValue <- "DOx_Hand_x_7"
   Button "Button_22" at 438,201 size 60x20; TextOff 'Вкл'; Authorization "Operate"
      on Click: SetBit("DOx_Start_M_x_7")
      Appearance <- "DOx_Start_M_x_7"
   Button "Button_23" at 548,225 size 20x20; TextOff 'Text'; Authorization "User administration"; PictureList "ok_green"
      on Click: InvertBit("DOx_Inverse_x_7")
      ProcessValue <- "DOx_Inverse_x_7"
   TextField "Text field_22" at 437,221 size 91x23; Text 'Инверсия:'
   IOField "I/O field_11" at 480,245 size 30x24; Authorization "Developer"; FormatPattern 99
      ProcessValue <- "DOx_ADDR_Byte_x_7"
   IOField "I/O field_12" at 520,245 size 20x24; Authorization "Developer"; FormatPattern 9
      ProcessValue <- "DOx_ADDR_Bit_x_7"
   TextField "Text field_23" at 462,245 size 20x23; Text 'Q'
   TextField "Text field_24" at 509,245 size 13x23; Text '.'
   Button "Button_41" at 590,176 size 130x22; TextOff 'Авто'; Authorization "Operate"; TextList "Hand"
      on Click: InvertBit("DOx_Hand_x_8")
      Appearance <- "DOx_Hand_x_8"
      ProcessValue <- "DOx_Hand_x_8"
   Button "Button_43" at 590,201 size 60x20; TextOff 'Вкл'; Authorization "Operate"
      on Click: SetBit("DOx_Start_M_x_8")
      Appearance <- "DOx_Start_M_x_8"
   Button "Button_44" at 700,225 size 20x20; TextOff 'Text'; Authorization "User administration"; PictureList "ok_green"
      on Click: InvertBit("DOx_Inverse_x_8")
      ProcessValue <- "DOx_Inverse_x_8"
   TextField "Text field_42" at 589,221 size 91x23; Text 'Инверсия:'
   IOField "I/O field_21" at 632,245 size 30x24; Authorization "Developer"; FormatPattern 99
      ProcessValue <- "DOx_ADDR_Byte_x_8"
   IOField "I/O field_22" at 672,245 size 20x24; Authorization "Developer"; FormatPattern 9
      ProcessValue <- "DOx_ADDR_Bit_x_8"
   TextField "Text field_43" at 614,245 size 20x23; Text 'Q'
   TextField "Text field_44" at 661,245 size 13x23; Text '.'
   Button "Button_24" at 134,312 size 130x22; TextOff 'Авто'; Authorization "Operate"; TextList "Hand"
      on Click: InvertBit("DOx_Hand_x_9")
      Appearance <- "DOx_Hand_x_9"
      ProcessValue <- "DOx_Hand_x_9"
   Button "Button_27" at 134,337 size 60x20; TextOff 'Вкл'; Authorization "Operate"
      on Click: SetBit("DOx_Start_M_x_9")
      Appearance <- "DOx_Start_M_x_9"
   Button "Button_28" at 244,361 size 20x20; TextOff 'Text'; PictureList "ok_green"; Authorization "User administration"
      on Click: InvertBit("DOx_Inverse_x_9")
      ProcessValue <- "DOx_Inverse_x_9"
   TextField "Text field_18" at 133,357 size 91x23; Text 'Инверсия:'
   IOField "I/O field_9" at 176,381 size 30x24; Authorization "Developer"; FormatPattern 99
      ProcessValue <- "DOx_ADDR_Byte_x_9"
   IOField "I/O field_10" at 216,381 size 20x24; Authorization "Developer"; FormatPattern 9
      ProcessValue <- "DOx_ADDR_Bit_x_9"
   TextField "Text field_19" at 158,381 size 20x23; Text 'Q'
   TextField "Text field_20" at 205,381 size 13x23; Text '.'
   Button "Button_37" at 286,312 size 130x22; TextOff 'Авто'; Authorization "Operate"; TextList "Hand"
      on Click: InvertBit("DOx_Hand_x_10")
      Appearance <- "DOx_Hand_x_10"
      ProcessValue <- "DOx_Hand_x_10"
   Button "Button_39" at 286,337 size 60x20; TextOff 'Вкл'; Authorization "Operate"
      on Click: SetBit("DOx_Start_M_x_10")
      Appearance <- "DOx_Start_M_x_10"
   Button "Button_40" at 396,361 size 20x20; TextOff 'Text'; Authorization "User administration"; PictureList "ok_green"
      on Click: InvertBit("DOx_Inverse_x_10")
      ProcessValue <- "DOx_Inverse_x_10"
   TextField "Text field_26" at 285,357 size 91x23; Text 'Инверсия:'
   IOField "I/O field_13" at 328,381 size 30x24; Authorization "Developer"; FormatPattern 99
      ProcessValue <- "DOx_ADDR_Byte_x_10"
   IOField "I/O field_14" at 368,381 size 20x24; Authorization "Developer"; FormatPattern 9
      ProcessValue <- "DOx_ADDR_Bit_x_10"
   TextField "Text field_27" at 310,381 size 20x23; Text 'Q'
   TextField "Text field_28" at 357,381 size 13x23; Text '.'
   Button "Button_48" at 590,312 size 130x22; TextOff 'Авто'; Authorization "Operate"; TextList "Hand"
      on Click: InvertBit("DOx_Hand_x_12")
      Appearance <- "DOx_Hand_x_12"
      ProcessValue <- "DOx_Hand_x_12"
   Button "Button_50" at 590,337 size 60x20; TextOff 'Вкл'; Authorization "Operate"
      on Click: SetBit("DOx_Start_M_x_12")
      Appearance <- "DOx_Start_M_x_12"
   Button "Button_51" at 700,361 size 20x20; TextOff 'Text'; Authorization "User administration"; PictureList "ok_green"
      on Click: InvertBit("DOx_Inverse_x_12")
      ProcessValue <- "DOx_Inverse_x_12"
   TextField "Text field_45" at 589,357 size 91x23; Text 'Инверсия:'
   IOField "I/O field_23" at 632,381 size 30x24; Authorization "Developer"; FormatPattern 99
      ProcessValue <- "DOx_ADDR_Byte_x_12"
   IOField "I/O field_24" at 672,381 size 20x24; Authorization "Developer"; FormatPattern 9
      ProcessValue <- "DOx_ADDR_Bit_x_12"
   TextField "Text field_46" at 614,381 size 20x23; Text 'Q'
   TextField "Text field_47" at 661,381 size 13x23; Text '.'
   TextField "Text field_38" at 438,283 size 130x26; Text 'выход 11'
   Button "Button_45" at 438,312 size 130x22; TextOff 'Авто'; Authorization "Operate"; TextList "Hand"
      on Click: InvertBit("DOx_Hand_x_11")
      Appearance <- "DOx_Hand_x_11"
      ProcessValue <- "DOx_Hand_x_11"
   Button "Button_47" at 438,337 size 60x20; TextOff 'Вкл'; Authorization "Operate"
      on Click: SetBit("DOx_Start_M_x_11")
      Appearance <- "DOx_Start_M_x_11"
   Button "Button_52" at 548,361 size 20x20; TextOff 'Text'; PictureList "ok_green"; Authorization "User administration"
      on Click: InvertBit("DOx_Inverse_x_11")